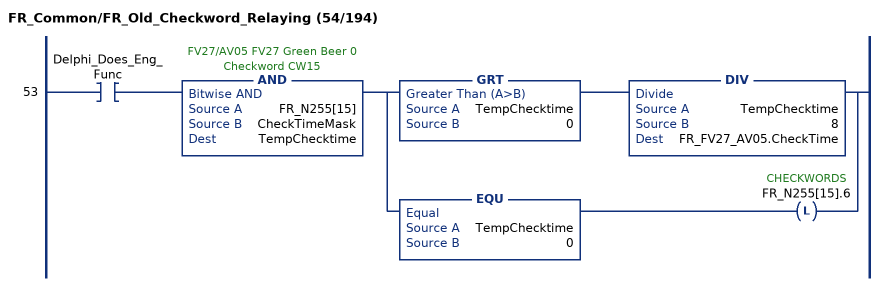
   53: XIC(Delphi_Does_Eng_Func)AND(FR_N255[15],CheckTimeMask,TempChecktime)[GRT(TempChecktime,0) DIV(TempChecktime,8,FR_FV27_AV05.CheckTime) ,EQU(TempChecktime,0) OTL(FR_N255[15].6) ];
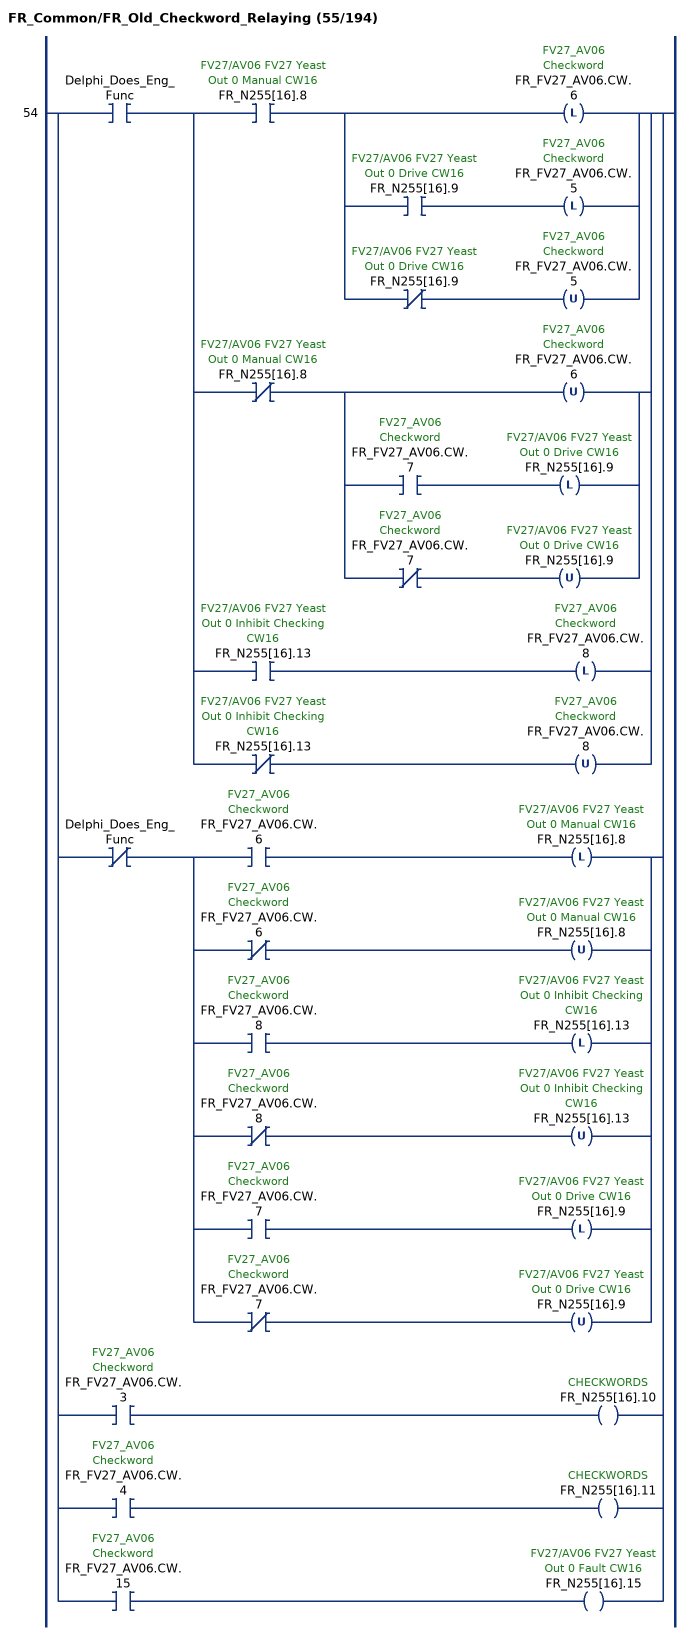
   54: [XIC(Delphi_Does_Eng_Func) [[XIC(FR_N255[16].8) [OTL(FR_FV27_AV06.CW.6) ,XIC(FR_N255[16].9) OTL(FR_FV27_AV06.CW.5) ,XIO(FR_N255[16].9) OTU(FR_FV27_AV06.CW.5) ] ,XIO(FR_N255[16].8) [OTU(FR_FV27_AV06.CW.6) ,[XIC(FR_FV27_AV06.CW.7) OTL(FR_N255[16].9) ,XIO(FR_FV27_AV06.CW.7) OTU(FR_N255[16].9) ] ] ] ,[XIC(FR_N255[16].13) OTL(FR_FV27_AV06.CW.8) ,XIO(FR_N255[16].13) OTU(FR_FV27_AV06.CW.8) ] ] ,XIO(Delphi_Does_Eng_Func) [[XIC(FR_FV27_AV06.CW.6) OTL(FR_N255[16].8) ,XIO(FR_FV27_AV06.CW.6) OTU(FR_N255[16].8) ] ,[XIC(FR_FV27_AV06.CW.8) OTL(FR_N255[16].13) ,XIO(FR_FV27_AV06.CW.8) OTU(FR_N255[16].13) ] ,[XIC(FR_FV27_AV06.CW.7) OTL(FR_N255[16].9) ,XIO(FR_FV27_AV06.CW.7) OTU(FR_N255[16].9) ] ] ,XIC(FR_FV27_AV06.CW.3) OTE(FR_N255[16].10) ,XIC(FR_FV27_AV06.CW.4) OTE(FR_N255[16].11) ,XIC(FR_FV27_AV06.CW.15) OTE(FR_N255[16].15) ];
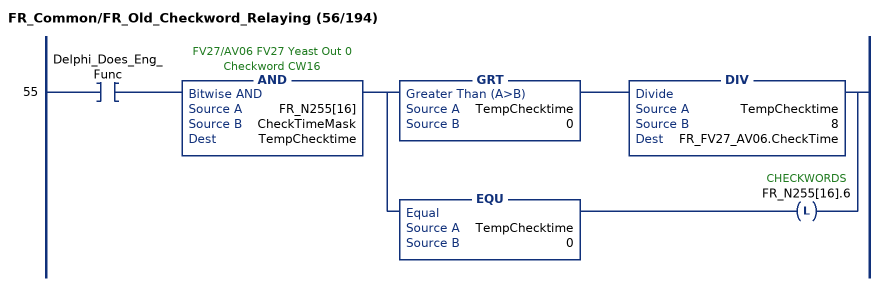
   55: XIC(Delphi_Does_Eng_Func)AND(FR_N255[16],CheckTimeMask,TempChecktime)[GRT(TempChecktime,0) DIV(TempChecktime,8,FR_FV27_AV06.CheckTime) ,EQU(TempChecktime,0) OTL(FR_N255[16].6) ];
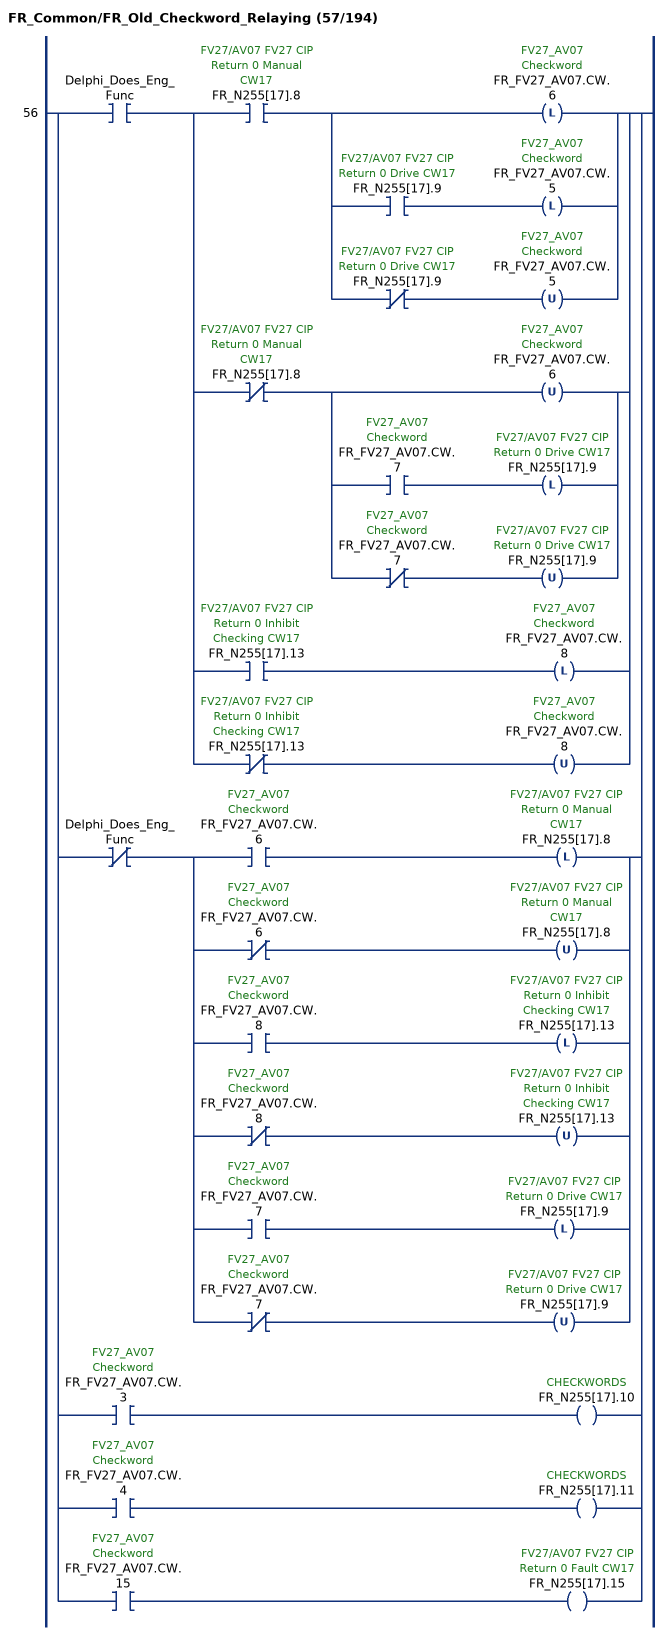
   56: [XIC(Delphi_Does_Eng_Func) [[XIC(FR_N255[17].8) [OTL(FR_FV27_AV07.CW.6) ,XIC(FR_N255[17].9) OTL(FR_FV27_AV07.CW.5) ,XIO(FR_N255[17].9) OTU(FR_FV27_AV07.CW.5) ] ,XIO(FR_N255[17].8) [OTU(FR_FV27_AV07.CW.6) ,[XIC(FR_FV27_AV07.CW.7) OTL(FR_N255[17].9) ,XIO(FR_FV27_AV07.CW.7) OTU(FR_N255[17].9) ] ] ] ,[XIC(FR_N255[17].13) OTL(FR_FV27_AV07.CW.8) ,XIO(FR_N255[17].13) OTU(FR_FV27_AV07.CW.8) ] ] ,XIO(Delphi_Does_Eng_Func) [[XIC(FR_FV27_AV07.CW.6) OTL(FR_N255[17].8) ,XIO(FR_FV27_AV07.CW.6) OTU(FR_N255[17].8) ] ,[XIC(FR_FV27_AV07.CW.8) OTL(FR_N255[17].13) ,XIO(FR_FV27_AV07.CW.8) OTU(FR_N255[17].13) ] ,[XIC(FR_FV27_AV07.CW.7) OTL(FR_N255[17].9) ,XIO(FR_FV27_AV07.CW.7) OTU(FR_N255[17].9) ] ] ,XIC(FR_FV27_AV07.CW.3) OTE(FR_N255[17].10) ,XIC(FR_FV27_AV07.CW.4) OTE(FR_N255[17].11) ,XIC(FR_FV27_AV07.CW.15) OTE(FR_N255[17].15) ];
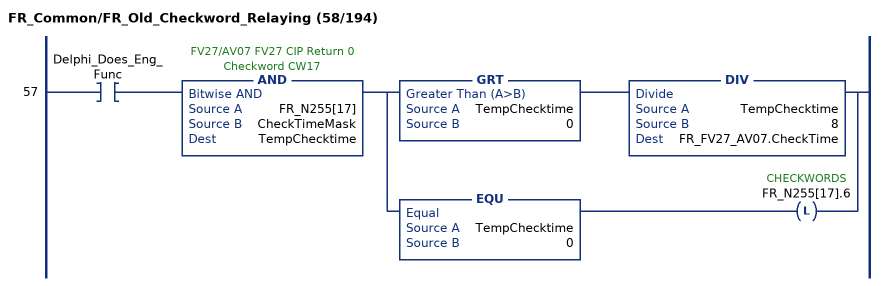
   57: XIC(Delphi_Does_Eng_Func)AND(FR_N255[17],CheckTimeMask,TempChecktime)[GRT(TempChecktime,0) DIV(TempChecktime,8,FR_FV27_AV07.CheckTime) ,EQU(TempChecktime,0) OTL(FR_N255[17].6) ];
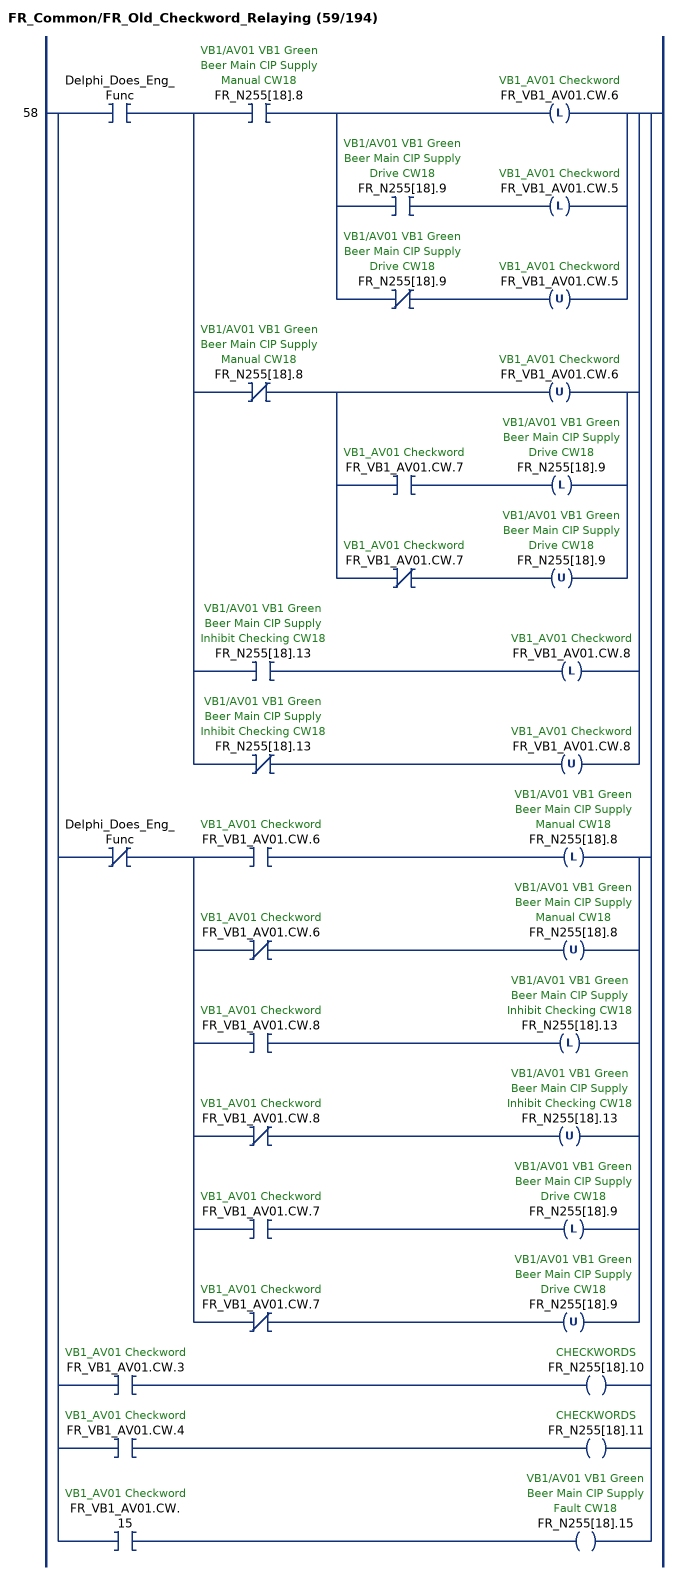
   58: [XIC(Delphi_Does_Eng_Func) [[XIC(FR_N255[18].8) [OTL(FR_VB1_AV01.CW.6) ,XIC(FR_N255[18].9) OTL(FR_VB1_AV01.CW.5) ,XIO(FR_N255[18].9) OTU(FR_VB1_AV01.CW.5) ] ,XIO(FR_N255[18].8) [OTU(FR_VB1_AV01.CW.6) ,[XIC(FR_VB1_AV01.CW.7) OTL(FR_N255[18].9) ,XIO(FR_VB1_AV01.CW.7) OTU(FR_N255[18].9) ] ] ] ,[XIC(FR_N255[18].13) OTL(FR_VB1_AV01.CW.8) ,XIO(FR_N255[18].13) OTU(FR_VB1_AV01.CW.8) ] ] ,XIO(Delphi_Does_Eng_Func) [[XIC(FR_VB1_AV01.CW.6) OTL(FR_N255[18].8) ,XIO(FR_VB1_AV01.CW.6) OTU(FR_N255[18].8) ] ,[XIC(FR_VB1_AV01.CW.8) OTL(FR_N255[18].13) ,XIO(FR_VB1_AV01.CW.8) OTU(FR_N255[18].13) ] ,[XIC(FR_VB1_AV01.CW.7) OTL(FR_N255[18].9) ,XIO(FR_VB1_AV01.CW.7) OTU(FR_N255[18].9) ] ] ,XIC(FR_VB1_AV01.CW.3) OTE(FR_N255[18].10) ,XIC(FR_VB1_AV01.CW.4) OTE(FR_N255[18].11) ,XIC(FR_VB1_AV01.CW.15) OTE(FR_N255[18].15) ];
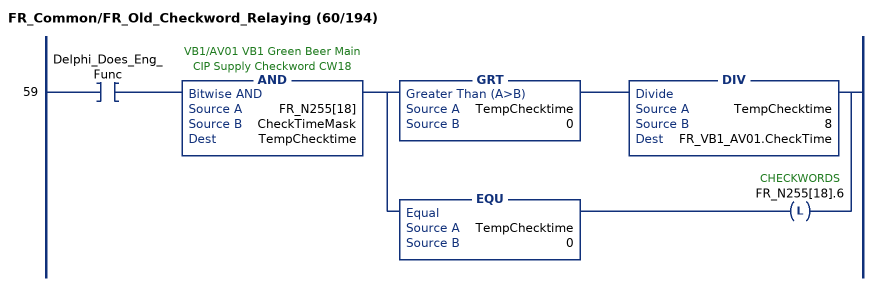
   59: XIC(Delphi_Does_Eng_Func)AND(FR_N255[18],CheckTimeMask,TempChecktime)[GRT(TempChecktime,0) DIV(TempChecktime,8,FR_VB1_AV01.CheckTime) ,EQU(TempChecktime,0) OTL(FR_N255[18].6) ];
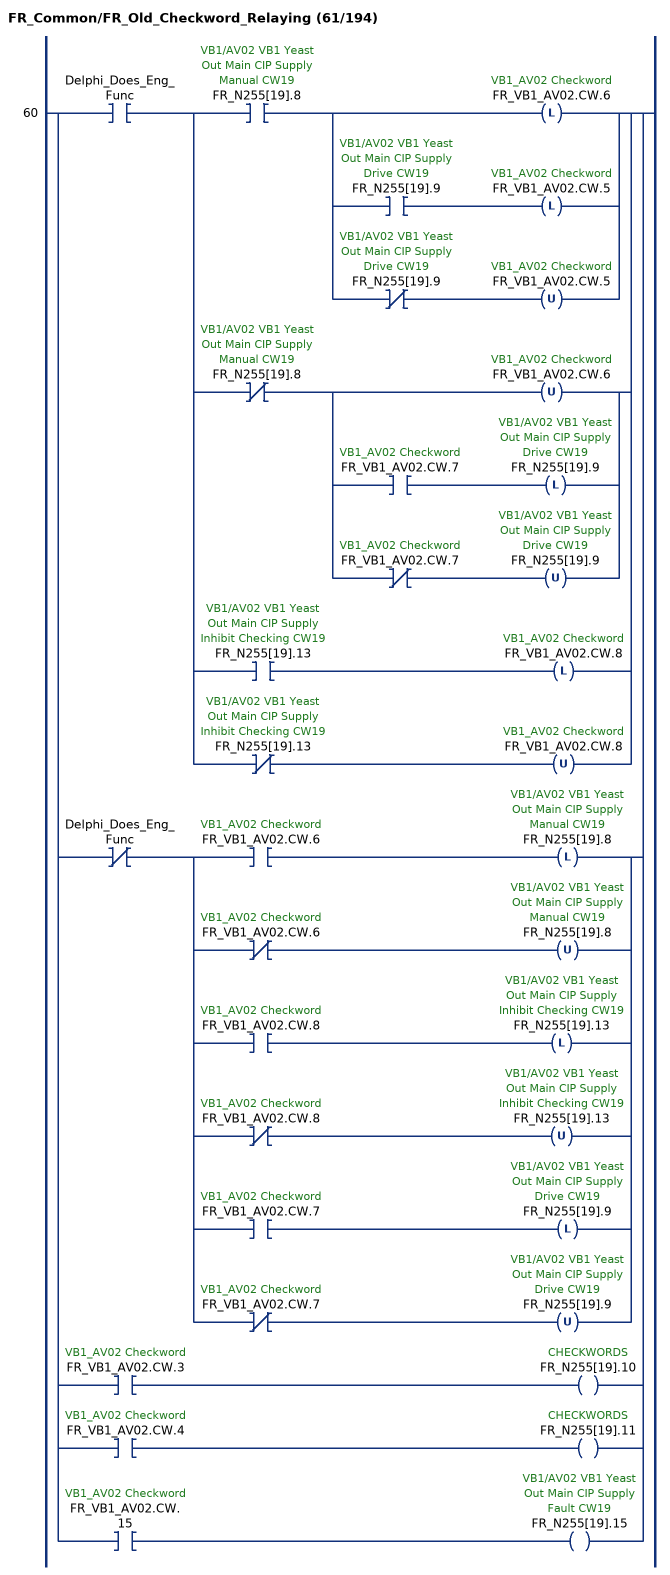
   60: [XIC(Delphi_Does_Eng_Func) [[XIC(FR_N255[19].8) [OTL(FR_VB1_AV02.CW.6) ,XIC(FR_N255[19].9) OTL(FR_VB1_AV02.CW.5) ,XIO(FR_N255[19].9) OTU(FR_VB1_AV02.CW.5) ] ,XIO(FR_N255[19].8) [OTU(FR_VB1_AV02.CW.6) ,[XIC(FR_VB1_AV02.CW.7) OTL(FR_N255[19].9) ,XIO(FR_VB1_AV02.CW.7) OTU(FR_N255[19].9) ] ] ] ,[XIC(FR_N255[19].13) OTL(FR_VB1_AV02.CW.8) ,XIO(FR_N255[19].13) OTU(FR_VB1_AV02.CW.8) ] ] ,XIO(Delphi_Does_Eng_Func) [[XIC(FR_VB1_AV02.CW.6) OTL(FR_N255[19].8) ,XIO(FR_VB1_AV02.CW.6) OTU(FR_N255[19].8) ] ,[XIC(FR_VB1_AV02.CW.8) OTL(FR_N255[19].13) ,XIO(FR_VB1_AV02.CW.8) OTU(FR_N255[19].13) ] ,[XIC(FR_VB1_AV02.CW.7) OTL(FR_N255[19].9) ,XIO(FR_VB1_AV02.CW.7) OTU(FR_N255[19].9) ] ] ,XIC(FR_VB1_AV02.CW.3) OTE(FR_N255[19].10) ,XIC(FR_VB1_AV02.CW.4) OTE(FR_N255[19].11) ,XIC(FR_VB1_AV02.CW.15) OTE(FR_N255[19].15) ];
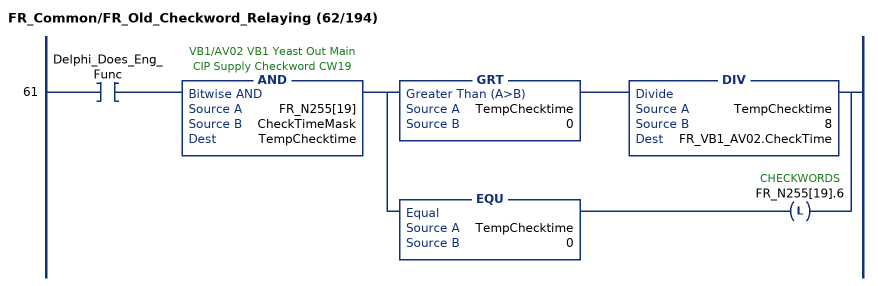
   61: XIC(Delphi_Does_Eng_Func)AND(FR_N255[19],CheckTimeMask,TempChecktime)[GRT(TempChecktime,0) DIV(TempChecktime,8,FR_VB1_AV02.CheckTime) ,EQU(TempChecktime,0) OTL(FR_N255[19].6) ];
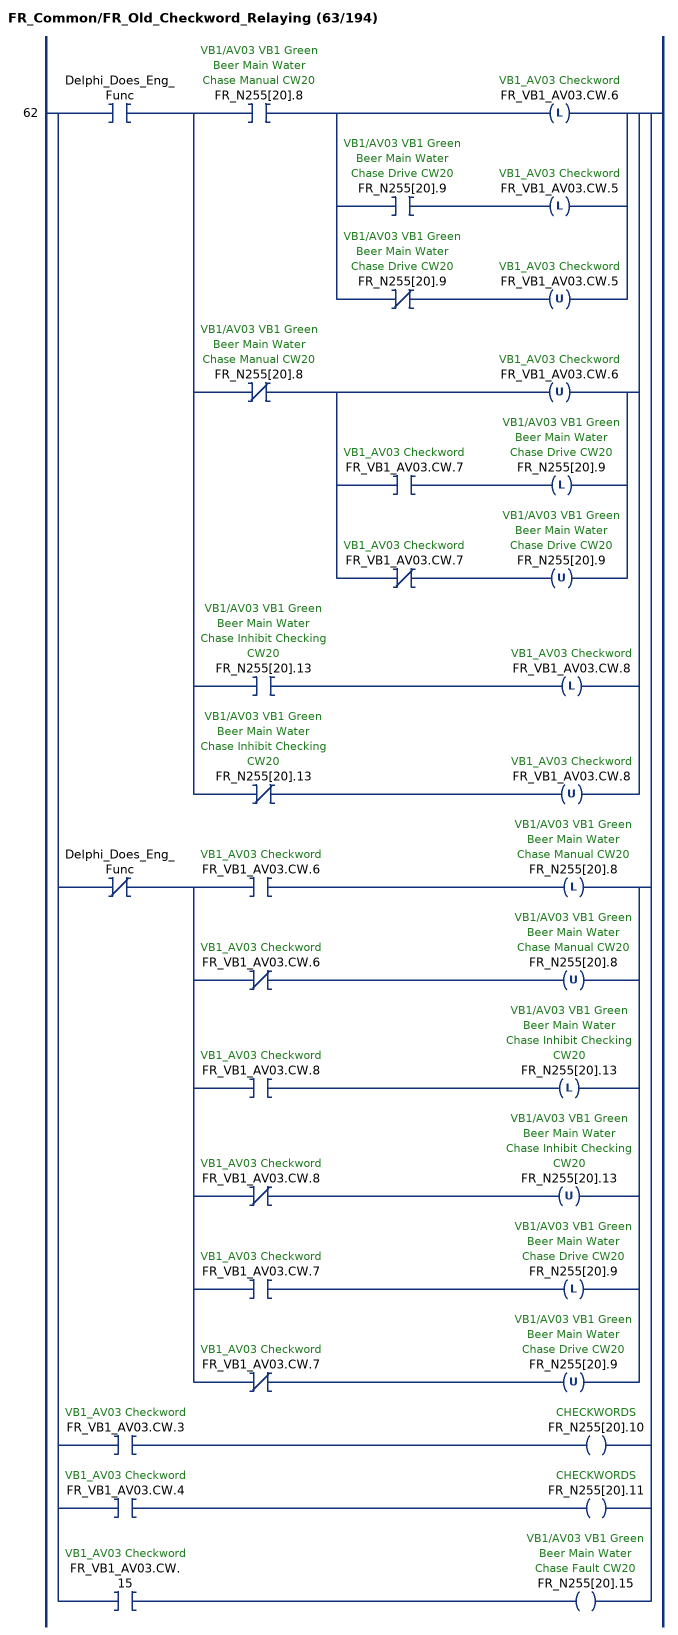
   62: [XIC(Delphi_Does_Eng_Func) [[XIC(FR_N255[20].8) [OTL(FR_VB1_AV03.CW.6) ,XIC(FR_N255[20].9) OTL(FR_VB1_AV03.CW.5) ,XIO(FR_N255[20].9) OTU(FR_VB1_AV03.CW.5) ] ,XIO(FR_N255[20].8) [OTU(FR_VB1_AV03.CW.6) ,[XIC(FR_VB1_AV03.CW.7) OTL(FR_N255[20].9) ,XIO(FR_VB1_AV03.CW.7) OTU(FR_N255[20].9) ] ] ] ,[XIC(FR_N255[20].13) OTL(FR_VB1_AV03.CW.8) ,XIO(FR_N255[20].13) OTU(FR_VB1_AV03.CW.8) ] ] ,XIO(Delphi_Does_Eng_Func) [[XIC(FR_VB1_AV03.CW.6) OTL(FR_N255[20].8) ,XIO(FR_VB1_AV03.CW.6) OTU(FR_N255[20].8) ] ,[XIC(FR_VB1_AV03.CW.8) OTL(FR_N255[20].13) ,XIO(FR_VB1_AV03.CW.8) OTU(FR_N255[20].13) ] ,[XIC(FR_VB1_AV03.CW.7) OTL(FR_N255[20].9) ,XIO(FR_VB1_AV03.CW.7) OTU(FR_N255[20].9) ] ] ,XIC(FR_VB1_AV03.CW.3) OTE(FR_N255[20].10) ,XIC(FR_VB1_AV03.CW.4) OTE(FR_N255[20].11) ,XIC(FR_VB1_AV03.CW.15) OTE(FR_N255[20].15) ];
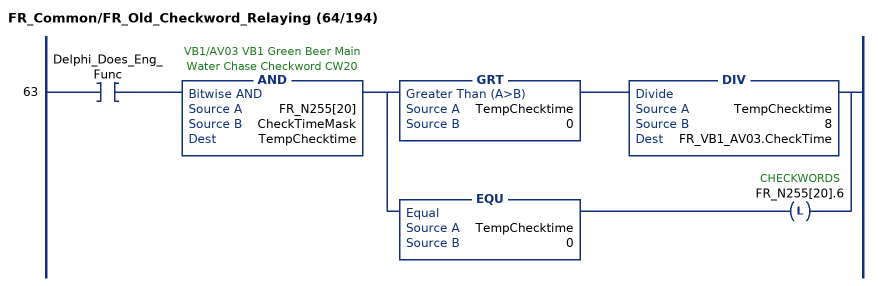
   63: XIC(Delphi_Does_Eng_Func)AND(FR_N255[20],CheckTimeMask,TempChecktime)[GRT(TempChecktime,0) DIV(TempChecktime,8,FR_VB1_AV03.CheckTime) ,EQU(TempChecktime,0) OTL(FR_N255[20].6) ];
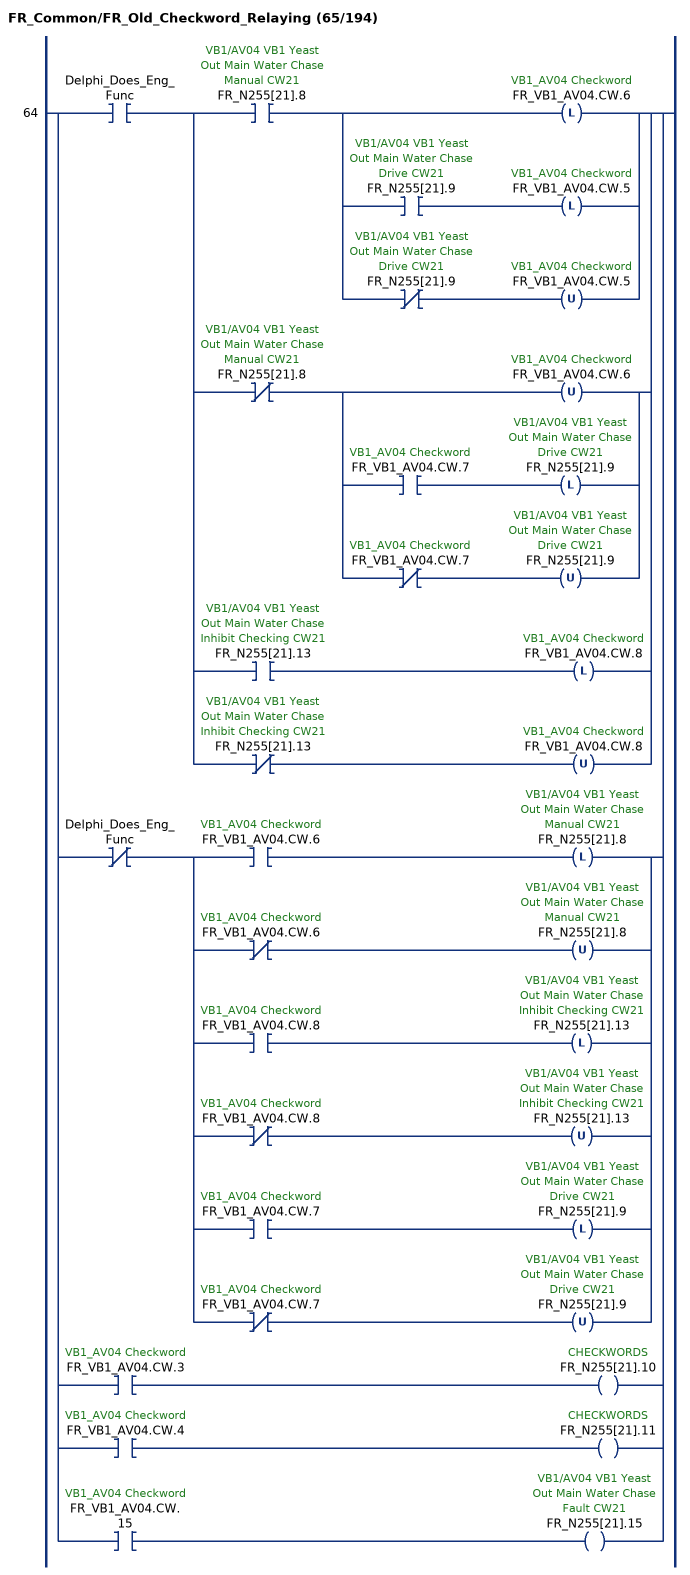
   64: [XIC(Delphi_Does_Eng_Func) [[XIC(FR_N255[21].8) [OTL(FR_VB1_AV04.CW.6) ,XIC(FR_N255[21].9) OTL(FR_VB1_AV04.CW.5) ,XIO(FR_N255[21].9) OTU(FR_VB1_AV04.CW.5) ] ,XIO(FR_N255[21].8) [OTU(FR_VB1_AV04.CW.6) ,[XIC(FR_VB1_AV04.CW.7) OTL(FR_N255[21].9) ,XIO(FR_VB1_AV04.CW.7) OTU(FR_N255[21].9) ] ] ] ,[XIC(FR_N255[21].13) OTL(FR_VB1_AV04.CW.8) ,XIO(FR_N255[21].13) OTU(FR_VB1_AV04.CW.8) ] ] ,XIO(Delphi_Does_Eng_Func) [[XIC(FR_VB1_AV04.CW.6) OTL(FR_N255[21].8) ,XIO(FR_VB1_AV04.CW.6) OTU(FR_N255[21].8) ] ,[XIC(FR_VB1_AV04.CW.8) OTL(FR_N255[21].13) ,XIO(FR_VB1_AV04.CW.8) OTU(FR_N255[21].13) ] ,[XIC(FR_VB1_AV04.CW.7) OTL(FR_N255[21].9) ,XIO(FR_VB1_AV04.CW.7) OTU(FR_N255[21].9) ] ] ,XIC(FR_VB1_AV04.CW.3) OTE(FR_N255[21].10) ,XIC(FR_VB1_AV04.CW.4) OTE(FR_N255[21].11) ,XIC(FR_VB1_AV04.CW.15) OTE(FR_N255[21].15) ];
